   //__________________________________________________________________
   // Shotcounter mixinghead 08:
   //
         A     "DB619_State_MPart".Mixinghead[1].Shotcounter."08";
         =     "DB123_MH_IO_Signals".MH[8].OUT.MH.H_Shotcounter_MH;
         JCN   countMH8end;
   //
         A     "DB619_State_MPart".Mixinghead[1].ImpCounterOn;
         JCN   countMH8end;
   //-----
         L     "DB_Zaehler_Anzeige".MH_Counter_Reset[8];
         L     "DB619_State_MPart".Mixinghead[1].Countervalue;
         DTR;
         +R;
         T     "DB_Zaehler_Anzeige".MH_Counter_Reset[8];
   //-----
         L     "DB_Zaehler_Anzeige".MH_Counter_NonReset[8];
         L     "DB619_State_MPart".Mixinghead[1].Countervalue;
         DTR;
         +R;
         T     "DB_Zaehler_Anzeige".MH_Counter_NonReset[8];
   //-----
         L     "DB_Zaehler_Schicht_aktuell".MH_Counter[8];
         L     1.0;
         +R;
         T     "DB_Zaehler_Schicht_aktuell".MH_Counter[8];
   //-----
   countMH8end:NOP   0;
   //__________________________________________________________________
   // Shotcounter mixinghead 09:
   //
         A     "DB619_State_MPart".Mixinghead[1].Shotcounter."09";
         =     "DB123_MH_IO_Signals".MH[9].OUT.MH.H_Shotcounter_MH;
         JCN   countMH9end;
   //
         A     "DB619_State_MPart".Mixinghead[1].ImpCounterOn;
         JCN   countMH9end;
   //-----
         L     "DB_Zaehler_Anzeige".MH_Counter_Reset[9];
         L     "DB619_State_MPart".Mixinghead[1].Countervalue;
         DTR;
         +R;
         T     "DB_Zaehler_Anzeige".MH_Counter_Reset[9];
   //-----
         L     "DB_Zaehler_Anzeige".MH_Counter_NonReset[9];
         L     "DB619_State_MPart".Mixinghead[1].Countervalue;
         DTR;
         +R;
         T     "DB_Zaehler_Anzeige".MH_Counter_NonReset[9];
   //-----
         L     "DB_Zaehler_Schicht_aktuell".MH_Counter[9];
         L     1.0;
         +R;
         T     "DB_Zaehler_Schicht_aktuell".MH_Counter[9];
   //-----
   countMH9end:NOP   0;
   //__________________________________________________________________
   // Shotcounter mixinghead 10:
   //
         A     "DB619_State_MPart".Mixinghead[1].Shotcounter."10";
         =     "DB123_MH_IO_Signals".MH[10].OUT.MH.H_Shotcounter_MH;
         JCN   countMH10end;
   //
         A     "DB619_State_MPart".Mixinghead[1].ImpCounterOn;
         JCN   countMH10end;
   //-----
         L     "DB_Zaehler_Anzeige".MH_Counter_Reset[10];
         L     "DB619_State_MPart".Mixinghead[1].Countervalue;
         DTR;
         +R;
         T     "DB_Zaehler_Anzeige".MH_Counter_Reset[10];
   //-----
         L     "DB_Zaehler_Anzeige".MH_Counter_NonReset[10];
         L     "DB619_State_MPart".Mixinghead[1].Countervalue;
         DTR;
         +R;
         T     "DB_Zaehler_Anzeige".MH_Counter_NonReset[10];
   //-----
         L     "DB_Zaehler_Schicht_aktuell".MH_Counter[10];
         L     1.0;
         +R;
         T     "DB_Zaehler_Schicht_aktuell".MH_Counter[10];
   //-----
   countMH10end:NOP   0;
END_REGION

REGION Network 8: Bits for nozzle/bypass control on mixinghead
         BEU;
   //______________________________________________________________
   // send nozzles for shot from shot data
         L;
         LAR1;
         L     "DB619_State_MPart".ShotMa[1].ShotData.Comp_at_Shot;
         T     LB[AR1, P#0.0];

         L;
         LAR1;
         L     "DB704_MH_Value".Mixinghead[1].NozzelCirc;
         T     LB[AR1, P#0.0];

         A     #TempNozzleShotConnection[1];
         AN    "DB753_MeteringPump".Pump[1].PumpDeselected;
         AN    "DB753_MeteringPump".Pump[1].PumpDeselectedInterval;
         =     #TempNozzleShotMH[1];
         =     #TempNozzleCirc[1];
         A     #TempNozzleShotConnection[2];
         AN    "DB753_MeteringPump".Pump[2].PumpDeselected;
         AN    "DB753_MeteringPump".Pump[2].PumpDeselectedInterval;
         =     #TempNozzleShotMH[2];
         =     #TempNozzleCirc[2];
         A     #TempNozzleShotConnection[3];
         AN    "DB753_MeteringPump".Pump[3].PumpDeselected;
         AN    "DB753_MeteringPump".Pump[3].PumpDeselectedInterval;
         =     #TempNozzleShotMH[3];
         =     #TempNozzleCirc[3];
         A     #TempNozzleShotConnection[4];
         AN    "DB753_MeteringPump".Pump[4].PumpDeselected;
         AN    "DB753_MeteringPump".Pump[4].PumpDeselectedInterval;
         =     #TempNozzleShotMH[4];
         =     #TempNozzleCirc[4];

         CLR;
         =     #TempNozzleShotMH[5];
         =     #TempNozzleCirc[5];

         L;
         LAR1;
         L     LB[AR1, P#0.0];
         T     "DB704_MH_Value".Mixinghead[1].NozzelShot;

   //______________________________________________________________
   // Nozzles in recirculation are different between cycle and recirculation
         AN    "DB619_State_MPart".Cycle[1].running;
         JC    rec;
         A     "DB619_State_MPart".Cycle[1].StandByTimeRuns;
         A     "DB619_State_MPart".Cycle[1].LastShotinToolFinished;
         AN    "DB619_State_MPart".ToolMa[1].ShotFound;
         AN    "DB619_State_MPart".Cycle[1].PulsShotend;
         S     #TempNozzleCirc[1];
         S     #TempNozzleCirc[2];
         S     #TempNozzleCirc[3];
         S     #TempNozzleCirc[4];
         JU    orec;
   rec:  A     "DB619_State_MPart".Recirculation[1].Lowpressure;
         JC    lopr;
         A     "DB619_State_MPart".Recirculation[1].Reduced;
         JC    rdpr;
         A     "DB619_State_MPart".Recirculation[1].Highpressure;
         JC    hdpr;
         JU    orec;

   // nozzles for lo pressure recirculation
   lopr: NOP   0;
         A     "DB704_MH_Value".Mixinghead[1].MH_Connection[1].LP_CircOverNozzle;
         =     #TempNozzleCirc[1];
         A     "DB704_MH_Value".Mixinghead[1].MH_Connection[2].LP_CircOverNozzle;
         =     #TempNozzleCirc[2];
         A     "DB704_MH_Value".Mixinghead[1].MH_Connection[3].LP_CircOverNozzle;
         =     #TempNozzleCirc[3];
         A     "DB704_MH_Value".Mixinghead[1].MH_Connection[4].LP_CircOverNozzle;
         =     #TempNozzleCirc[4];
         JU    orec;
   // nozzles for reduced recirculation
   rdpr: A     "DB704_MH_Value".Mixinghead[1].MH_Connection[1].Red_CircOverNozzle;
         =     #TempNozzleCirc[1];
         A     "DB704_MH_Value".Mixinghead[1].MH_Connection[2].Red_CircOverNozzle;
         =     #TempNozzleCirc[2];
         A     "DB704_MH_Value".Mixinghead[1].MH_Connection[3].Red_CircOverNozzle;
         =     #TempNozzleCirc[3];
         A     "DB704_MH_Value".Mixinghead[1].MH_Connection[4].Red_CircOverNozzle;
         =     #TempNozzleCirc[4];
         JU    orec;
   // nozzles for high pressure recirculation
   hdpr: A     "DB704_MH_Value".Mixinghead[1].MH_Connection[1].HP_CircOverNozzle;
         =     #TempNozzleCirc[1];
         A     "DB704_MH_Value".Mixinghead[1].MH_Connection[2].HP_CircOverNozzle;
         =     #TempNozzleCirc[2];
         A     "DB704_MH_Value".Mixinghead[1].MH_Connection[3].HP_CircOverNozzle;
         =     #TempNozzleCirc[3];
         A     "DB704_MH_Value".Mixinghead[1].MH_Connection[4].HP_CircOverNozzle;
         =     #TempNozzleCirc[4];
         JU    orec;

   // switch deselected components to bypass before sending info to procan module
   orec: NOP   0;
         O     "DB753_MeteringPump".Pump[1].PumpDeselected;
         O     "DB613_Komponent_State".MeteringPump[1].IntervalPause;
         R     #TempNozzleCirc[1];
         O     "DB753_MeteringPump".Pump[2].PumpDeselected;
         O     "DB613_Komponent_State".MeteringPump[2].IntervalPause;
         R     #TempNozzleCirc[2];
         O     "DB753_MeteringPump".Pump[3].PumpDeselected;
         O     "DB613_Komponent_State".MeteringPump[3].IntervalPause;
         R     #TempNozzleCirc[3];
         O     "DB753_MeteringPump".Pump[4].PumpDeselected;
         O     "DB613_Komponent_State".MeteringPump[4].IntervalPause;
         R     #TempNozzleCirc[4];

         A     "TM_SwitchOnDelayFCPump";
         JCN   PUND;
         SET;
         R     #TempNozzleCirc[1];
         R     #TempNozzleCirc[2];
         R     #TempNozzleCirc[3];
         R     #TempNozzleCirc[4];
         JU    NozC;

   PUND: O     "DB619_State_MPart".Recirculation[1].Lowpressure;
         O     "DB619_State_MPart".Recirculation[1].Reduced;
         AN    "DB619_State_MPart".Recirculation[1].Pausetime;
         O     "DB619_State_MPart".Recirculation[1].Highpressure;
         O     "DB619_State_MPart".Cycle[1].running;
         JCN   mask;

   NozC: NOP   0;

         L;
         LAR1;
         L     LB[AR1, P#0.0];
         T     "DB704_MH_Value".Mixinghead[1].NozzelCirc;

   //______________________________________________________________
   // Mask with enable bits for the nozzle/bypass pairs
   mask: L;
         LAR1;
         L     0;
         T     LW[AR1, P#0.0];

   // Jump over enabling of nozzles when nozzle leakage test is active
         A     "DB704_MH_Value".Mixinghead[1].NozzleLeakageTest;
         A     "DB619_State_MPart".Operationmode[1].Manual;
         JC    test;

         A     "DB613_Komponent_State".MeteringPump[1].Main_Pumpselection;
         =     #TempMask.EnableNozzle_1;
         A     "DB613_Komponent_State".MeteringPump[2].Main_Pumpselection;
         =     #TempMask.EnableNozzle_2;
         A     "DB613_Komponent_State".MeteringPump[3].Main_Pumpselection;
         =     #TempMask.EnableNozzle_3;
         A     "DB613_Komponent_State".MeteringPump[4].Main_Pumpselection;
         =     #TempMask.EnableNozzle_4;

   test: L;
         LAR1;

         L     LW[AR1, P#0.0];  // target status
         L     "DB704_MH_Value".Mixinghead[1].NozzelForcen;  // old status
         XOW;  //  -> bits with differences
         AW;  // compare again with accu 2 -> bits to be switched on
         T     #SwitchOn;

         L     "DB704_MH_Value".Mixinghead[1].NozzelForcen;  // old status
         L     LW[AR1, P#0.0];  // target status
         XOW;  // -> bits with differences
         AW;  // compare again with accu 2 -> bits to be switched off
         T     #SwitchOff;

         A     <>0;
         L     "DB704_MH_Value".Mixinghead[1].DelayTimeNozzlesOff;
         SD    "TM_Nozzle_off_delay_MH01";
         A     "TM_Nozzle_off_delay_MH01";
         JCN   nzon;
         L     "DB704_MH_Value".Mixinghead[1].NozzelForcen;
         L     #SwitchOff;
         XOW;
         T     "DB704_MH_Value".Mixinghead[1].NozzelForcen;

   nzon: L     #SwitchOn;
         L     "DB704_MH_Value".Mixinghead[1].NozzelForcen;
         OW;
         T     "DB704_MH_Value".Mixinghead[1].NozzelForcen;

         A     "DB704_MH_Value".Mixinghead[1].NozzleLeakageTest;
         =     "DB824_Error_MH_CP".MH_Control[0].WRN_NozzleLeakageTest_active;
END_REGION
END_FUNCTION_BLOCK

FUNCTION_BLOCK "FB015_MeteringPump_M1"   // FB15, STL
TITLE = Meteringunit, edge filter, feed pump
{ S7_Optimized_Access := 'FALSE' }
AUTHOR : KT242
VERSION : 0.1
// Control of metering unit
   VAR_TEMP
      Dummy : Bool;
      Release_external : Bool;
      Release_FU : Bool;
      active : Bool;
      High_speed : Bool;
      V_2_Point_adjustment : Bool;
      Imp_WT_Ein : Bool;
      Imp_WT_Aus : Bool;
      HM_Intervall_Aus : Bool;
      Temp_F_FU_Poly : Bool;
      Temp_F_FU_Iso : Bool;
      Temp_enableCL_k1 : Bool;
      Temp_enableCL_k2 : Bool;
      Temp_Enable_C1 : Bool;
      Temp_Press_OK : Bool;
      CompUsedForShot : Array[1..16] of Bool;
      RetValSFC : Int;
   END_VAR
BEGIN

REGION Network 1: Min.- and Max.-value pump

         CALL  "FC217_Calc_flow_limits";
END_REGION

REGION Network 2

         CALL  "FC051_ComponentGeneral";
END_REGION

REGION Network 3: Temperautre control

         CALL  "FC057_HPHeatexchanger";
         CALL  "FC057_LPHeatexchanger";
END_REGION

REGION Network 4: Switch ON delay FU pump
   //-----
         O(;
         AN    "DB619_State_MPart".Machine[1].Metering."01";
         AN    "DB753_MeteringPump".Pump[1].PumpDeselected;
         A     "DB753_MeteringPump".Pump[1].WithFC;
         );
         O(;
         AN    "DB619_State_MPart".Machine[1].Metering."02";
         AN    "DB753_MeteringPump".Pump[2].PumpDeselected;
         A     "DB753_MeteringPump".Pump[2].WithFC;
         );
         O(;
         AN    "DB619_State_MPart".Machine[1].Metering."03";
         AN    "DB753_MeteringPump".Pump[3].PumpDeselected;
         A     "DB753_MeteringPump".Pump[3].WithFC;
         );
         O(;
         AN    "DB619_State_MPart".Machine[1].Metering."04";
         AN    "DB753_MeteringPump".Pump[4].PumpDeselected;
         A     "DB753_MeteringPump".Pump[4].WithFC;
         );
         O(;
         AN    "DB619_State_MPart".Machine[1].Metering."05";
         AN    "DB753_MeteringPump".Pump[5].PumpDeselected;
         A     "DB753_MeteringPump".Pump[5].WithFC;
         );
         O(;
         AN    "DB619_State_MPart".Machine[1].Metering."06";
         AN    "DB753_MeteringPump".Pump[6].PumpDeselected;
         A     "DB753_MeteringPump".Pump[6].WithFC;
         );
         FP    "HF_FP_SwitchOffPump";
         =     "PulsePumpSwitchedOff";
         L     S5T#5S;
         SE    "TM_SwitchOnDelayFCPump";
   //-----
END_REGION

REGION Network 5: Release of pumps
   // Copy Control bits for module to local area
         L;
         LAR1;
         L     "DB619_State_MPart".ShotMa[1].ShotData.Comp_at_Shot;
         CAW;
         T     LW[AR1, P#0.0];
   //-----
         A(;
         O     "DB619_State_MPart".CylinderManager[1].Selection_Metering;
         ON    "DB619_State_MPart".CylinderManager[1].Block_is_active;
         );
   //-----
         A(;
         O     "DB613_Komponent_State".MeteringPump[1].Main_Pumpselection;
         O     "DB753_MeteringPump".Pump[1].PumpDeselected;
         O     "DB613_Komponent_State".MeteringPump[1].IntervalPause;
         ON    "DB613_Komponent_State".MeteringPump[1].Block_is_active;
         );
         A(;
         O     "DB613_Komponent_State".MeteringPump[2].Main_Pumpselection;
         O     "DB753_MeteringPump".Pump[2].PumpDeselected;
         O     "DB613_Komponent_State".MeteringPump[2].IntervalPause;
         ON    "DB613_Komponent_State".MeteringPump[2].Block_is_active;
         );
         A(;
         O     "DB613_Komponent_State".MeteringPump[3].Main_Pumpselection;
         O     "DB753_MeteringPump".Pump[3].PumpDeselected;
         O     "DB613_Komponent_State".MeteringPump[3].IntervalPause;
         ON    "DB613_Komponent_State".MeteringPump[3].Block_is_active;
         );
         A(;
         O     "DB613_Komponent_State".MeteringPump[4].Main_Pumpselection;
         O     "DB753_MeteringPump".Pump[4].PumpDeselected;
         O     "DB613_Komponent_State".MeteringPump[4].IntervalPause;
         ON    "DB613_Komponent_State".MeteringPump[4].Block_is_active;
         );
         A(;
         O     "DB613_Komponent_State".MeteringPump[5].Main_Pumpselection;
         O     "DB753_MeteringPump".Pump[5].PumpDeselected;
         O     "DB613_Komponent_State".MeteringPump[5].IntervalPause;
         ON    "DB613_Komponent_State".MeteringPump[5].Block_is_active;
         );
         A(;
         O     "DB613_Komponent_State".MeteringPump[6].Main_Pumpselection;
         O     "DB753_MeteringPump".Pump[6].PumpDeselected;
         O     "DB613_Komponent_State".MeteringPump[6].IntervalPause;
         ON    "DB613_Komponent_State".MeteringPump[6].Block_is_active;
         );
         AN    "TM_SwitchOnDelayFCPump";
         AN    "TM_Interrupt2PointAdjustment";
         =     #Release_external;
   //-----
END_REGION

REGION Network 6: Preparation for 2 Point- Adjustment
         CALL  "FC216_2-point_adjust";
END_REGION

REGION Network 7: Component 1
   //___________________________________________________________________________
   // Feedpump component 1
   //___________________________________________________________________________
   //
         CALL  "FC123_FeedingPump"
         ( IN_Release               := "DB619_State_MPart".Operationmode[1].valid,
           IN_ControlVoltage        := "DB619_State_MPart".Operationmode[1].Controllvoltage,
           IN_Reset_fault           := "DB009_Faults".Faults_Reset_FKT_M1,
           IN_ComponentDeselected   := "DB613_Komponent_State".MeteringPump[1].Mes_PumpDeselected,
           IN_Request_Feed          := "DB613_Komponent_State".MeteringPump[1].Selection_Feedingpump,
           IN_Request_Filling       := "DB612_Tank_State".Tank[1].Filling_Start,
           IN_Request_Bypass        := 1,
           IN_Fault_Motorprotection := "F_FeedingP_C1",
           IN_FaultFreqConverter    := "F_FCFeedingP_C1",
           IN_DryRun                := "DB612_Tank_State".Tank[1].Min_Level,
           IN_MaxLevelTray          := "DB612_Tank_State".Tank[1].LevelTriptray,
           IN_MaxPressure           := 1,
           IN_TempRelease           := 1,
           IN_TimerDrive            := "TM1_FeedPump01",
           IN_TimerStartUpFConv     := "TM2_FeedPump01",
           Values                   := "DB751_auxiliaryDriveMetering".FeedingPump[1],
           OUT_MainsContactor       := "M_FeedingP_C1",
           OUT_Release_FConverter   := "M_FeedingP_Start_C1",
           IO_Status                := "DB613_Komponent_State".FeedPump[1],
           IO_NewFault              := "DB009_Faults".Faultschanging_M1,
           IO_FaultLevel_1          := "DB009_Faults".Faults_FKT_Grp_1_M1,
           IO_FaultLevel_3          := "DB009_Faults".Faults_FKT_Grp_3_M1,
           IO_Faults                := "DB823_Error_Metering".FeedPump[1]
         );
   //___________________________________________________________________________
   // Edgefilter component 1
   //___________________________________________________________________________
   //
         CALL  "FC122_EdgeFilter"
         ( IN_Release               := "DB619_State_MPart".Operationmode[1].valid,
           IN_Reset_fault           := "DB009_Faults".Faults_Reset_FKT_M1,
           IN_Fault_Motorprotection := "F_Platefilter_C1",
           IN_DifPressure           := FALSE,
           IN_TimerDrive            := "TM_EdgeFilter01",
           Values                   := "DB751_auxiliaryDriveMetering".EdgeFilter[1],
           OUT_MainsContactor       := "M_Platefilter_C1",
           IO_Status                := "DB613_Komponent_State".EdgeFilter[1],
           IO_NewFault              := "DB009_Faults".Faultschanging_M1,
           IO_FaultLevel_3          := "DB009_Faults".Faults_FKT_Grp_3_M1,
           IO_Faults                := "DB823_Error_Metering".EdgeFilter[1]
         );
   //___________________________________________________________________________
   // Metering pump component 1
   //___________________________________________________________________________
   //
         A     "P_Min_C1";
         O;
         A     "DB619_State_MPart".Operationmode[1].Test;
         A     "V_Bypass_C1";
         =     #Temp_Press_OK;

         O     "DB612_Tank_State".Pentan[1].EnableComponentPump;
         ON    "DB702_Tank_Value".Tank[1].With_Filling_Pentane;
         A     #Release_external;
         =     #Temp_Enable_C1;
   //-----
         CALL  "FC053_MeteringPump"
         ( IN_ControlVoltage        := "DB619_State_MPart".Operationmode[1].Controllvoltage,
           IN_OperationMode_Valid   := #Release_external,
           IN_OPerationMode_Active  := "DB619_State_MPart".Operationmode[1].Active,
           IN_Min_PrePressure       := "P_Prepressure_Pump_C1",
           IN_Max_PressureComponent := "P_Max_C1",
           IN_MotorprotectionPump   := "F_Pump_C1",
           IN_With_FU_Pump          := "DB753_MeteringPump".Pump[1].WithFC,
           IN_FLT_FU_Pump           := "F_FC_Pump_C1",
           IN_MaxLevelTray          := "L_DripTray_C1",
           IN_Shot_Start            := "DB619_State_MPart".Cycle[1].Shotrelease,
           IN_MinPressure           := #Temp_Press_OK,  //"P_Min_C1"
           IN_PreAlarmBearing       := FALSE,  // "F_PreAlarmBearing_K2"
           IN_AlarmBearing          := FALSE,  // "F_AlarmBearing_K2"
           IN_Reset_fault_Fkt       := "DB009_Faults".Faults_Reset_FKT_M1,
           IN_ReleaseExternal       := #Temp_Enable_C1,  // #Release_external
           IN_FaultGroup_1          := "DB009_Faults".Fault_State_Grp_1_M1,
           IN_SOverSOffSWU_running  := "DB619_State_MPart".SWU[1].Switchingtime_runs,
           IN_High_speed            := 0,
           IN_2point_Adjustment     := "DB613_Komponent_State".MeteringPump[1]."2PointAdjustmentSelected",
           IN_Cycle_running         := "DB619_State_MPart".Cycle[1].running,
           IN_Recirc_reduced        := "DB619_State_MPart".Recirculation[1].Reduced,
           IN_Recirc_lowpressure    := "DB619_State_MPart".Recirculation[1].Lowpressure,
           IN_Recirc_highpressure   := "DB619_State_MPart".Recirculation[1].Highpressure,
           IN_Recirc_pausetime      := "DB619_State_MPart".Recirculation[1].Pausetime,
           IN_UsedForShot           := #CompUsedForShot[1],
           IN_Delay_Restart         := S5T#2S,
           IN_Timer_Restart         := "TM_RestartC01",
           IN_RunDownTime_FeedPump  := S5T#3S,
           IN_Timer_ControlFeedPump := "TM_CtrlFeedPumpC01",
           IN_TimerOffFeedPump      := "TM_CommonC01",
           IN_Timer_Delay_EnClosedL := "TM_DelayClosedLoopC01",
           IN_TimerInterval         := "TM_IntervalC01",
           OUT_2_Point_Adjust       := #V_2_Point_adjustment,
           OUT_Dosing_active        := #Dummy,
           OUT_Enableclosedloop     := "DB122_FlowIndexState".MeteringUnit[1].OUT_PROCAN.FlowIndex.Enableclosedloop,
           OUT_Pump_MainsContactor  := "M_Pump_Net_C1",
           OUT_Release_FU           := "M_Pump_Start_C1",
           IO_QPB_Pumpe             := "DB122_FlowIndexState".MeteringUnit[1].OUT_PROCAN.FlowIndex.StartQPB,
           IO_Status                := "DB613_Komponent_State".MeteringPump[1],
           IO_Fault                 := "DB823_Error_Metering".MeteringPump[1],
           IO_Config                := "DB753_MeteringPump".Pump[1],
           IO_NewFault              := "DB009_Faults".Faultschanging_M1,
           IO_FaultLevel_1          := "DB009_Faults".Faults_FKT_Grp_1_M1,
           IO_FaultLevel_2          := "DB009_Faults".Faults_FKT_Grp_2_M1,
           IO_FaultLevel_3          := "DB009_Faults".Faults_FKT_Grp_3_M1
         );
   //-----
   //-----
   // 2 Point adjustment
         A     #V_2_Point_adjustment;
         L     s5t#800ms;
         SE    "TM_pulse_2PointAdjust_C1";

         A     #V_2_Point_adjustment;
         L     s5t#500ms;
         SD    "TM_delay_2PointAdjust_C1";
         A     "TM_delay_2PointAdjust_C1";
         =     "V_Pump_2Point_C1";
   //-----
   //
         A     "DB613_Komponent_State".MeteringPump[1].Metering_to_PUC;
         =     "DB619_State_MPart".Machine[1].Metering."01";
   //
         A     "DB613_Komponent_State".MeteringPump[1].Metering_to_PUC;
         =     "M1C01active";
   //___________________________________________________________________________
   // Ventilation metering pump component 1
   //___________________________________________________________________________
   //
         CALL  "FC055_PumpVentilation"
         ( IN_Reset_fault_Fkt     := "DB009_Faults".Faults_Reset_FKT_M1,
           IN_Motorprotection     := "F_Fan_Pump_C1",
           IN_ComponentDeselected := "DB613_Komponent_State".MeteringPump[1].Mes_PumpDeselected,
           In_Start               := "DB613_Komponent_State".MeteringPump[1].Metering_to_PUC,
           IN_Time                := S5T#1M,
           IN_Timer               := "TM_FanPumpC01",
           OUT_MainContactor      := "M_Fan_Pump_Net_C1",
           IO_FLT_MotorFan        := "DB823_Error_Metering".MeteringPump[1].FLT_MotorFan,
           IO_NewFault            := "DB009_Faults".Faultschanging_M1,
           IO_FaultLevel_2        := "DB009_Faults".Faults_FKT_Grp_2_M1,
           IO_FaultLevel_3        := "DB009_Faults".Faults_FKT_Grp_3_M1
         );
   //
END_REGION

REGION Network 8: Component 2
   //___________________________________________________________________________
   // Feedpump component 2
   //___________________________________________________________________________
   //
         CALL  "FC123_FeedingPump"
         ( IN_Release               := "DB619_State_MPart".Operationmode[1].valid,
           IN_ControlVoltage        := "DB619_State_MPart".Operationmode[1].Controllvoltage,
           IN_Reset_fault           := "DB009_Faults".Faults_Reset_FKT_M1,
           IN_ComponentDeselected   := "DB613_Komponent_State".MeteringPump[2].Mes_PumpDeselected,
           IN_Request_Feed          := "DB613_Komponent_State".MeteringPump[2].Selection_Feedingpump,
           IN_Request_Filling       := 0,
           IN_Request_Bypass        := 0,
           IN_Fault_Motorprotection := "F_FeedingP_C2",
           IN_FaultFreqConverter    := "F_FCFeedingP_C2",
           IN_DryRun                := "DB612_Tank_State".Tank[2].Min_Level,
           IN_MaxLevelTray          := "DB612_Tank_State".Tank[2].LevelTriptray,
           IN_MaxPressure           := 1,
           IN_TempRelease           := 1,
           IN_TimerDrive            := "TM1_FeedPump02",
           IN_TimerStartUpFConv     := "TM2_FeedPump02",
           Values                   := "DB751_auxiliaryDriveMetering".FeedingPump[2],
           OUT_MainsContactor       := "M_FeedingP_C2",
           OUT_Release_FConverter   := "M_FeedingP_Start_C2",
           IO_Status                := "DB613_Komponent_State".FeedPump[2],
           IO_NewFault              := "DB009_Faults".Faultschanging_M1,
           IO_FaultLevel_1          := "DB009_Faults".Faults_FKT_Grp_1_M1,
           IO_FaultLevel_3          := "DB009_Faults".Faults_FKT_Grp_3_M1,
           IO_Faults                := "DB823_Error_Metering".FeedPump[2]
         );
   //___________________________________________________________________________
   // Edgefilter component 2
   //___________________________________________________________________________
   //
         CALL  "FC122_EdgeFilter"
         ( IN_Release               := "DB619_State_MPart".Operationmode[1].valid,
           IN_Reset_fault           := "DB009_Faults".Faults_Reset_FKT_M1,
           IN_Fault_Motorprotection := "F_Platefilter_C2",
           IN_DifPressure           := FALSE,
           IN_TimerDrive            := "TM_EdgeFilter02",
           Values                   := "DB751_auxiliaryDriveMetering".EdgeFilter[2],
           OUT_MainsContactor       := "M_Platefilter_C2",
           IO_Status                := "DB613_Komponent_State".EdgeFilter[2],
           IO_NewFault              := "DB009_Faults".Faultschanging_M1,
           IO_FaultLevel_3          := "DB009_Faults".Faults_FKT_Grp_3_M1,
           IO_Faults                := "DB823_Error_Metering".EdgeFilter[2]
         );
   //___________________________________________________________________________
   // Metering pump component 2
   //___________________________________________________________________________
   //
         A     "P_Min_C2";
         O;
         A     "DB619_State_MPart".Operationmode[1].Test;
         A     "V_Bypass_C2";
         =     #Temp_Press_OK;

         CALL  "FC053_MeteringPump"
         ( IN_ControlVoltage        := "DB619_State_MPart".Operationmode[1].Controllvoltage,
           IN_OperationMode_Valid   := #Release_external,  // not used at FC
           IN_OPerationMode_Active  := "DB619_State_MPart".Operationmode[1].Active,
           IN_Min_PrePressure       := "P_Prepressure_Pump_C2",
           IN_Max_PressureComponent := "P_Max_C2",
           IN_MotorprotectionPump   := "F_Pump_C2",
           IN_With_FU_Pump          := "DB753_MeteringPump".Pump[2].WithFC,
           IN_FLT_FU_Pump           := "F_FC_Pump_C2",
           IN_MaxLevelTray          := "L_DripTray_C2",
           IN_Shot_Start            := "DB619_State_MPart".Cycle[1].Shotrelease,
           IN_MinPressure           := #Temp_Press_OK,  //"P_Min_C2"
           IN_PreAlarmBearing       := FALSE,  // "F_PreAlarmBearing_K2"
           IN_AlarmBearing          := FALSE,  // "F_AlarmBearing_K2"
           IN_Reset_fault_Fkt       := "DB009_Faults".Faults_Reset_FKT_M1,
           IN_ReleaseExternal       := #Release_external,
           IN_FaultGroup_1          := "DB009_Faults".Fault_State_Grp_1_M1,
           IN_SOverSOffSWU_running  := "DB619_State_MPart".SWU[1].Switchingtime_runs,
           IN_High_speed            := 0,
           IN_2point_Adjustment     := "DB613_Komponent_State".MeteringPump[2]."2PointAdjustmentSelected",
           IN_Cycle_running         := "DB619_State_MPart".Cycle[1].running,
           IN_Recirc_reduced        := "DB619_State_MPart".Recirculation[1].Reduced,
           IN_Recirc_lowpressure    := "DB619_State_MPart".Recirculation[1].Lowpressure,
           IN_Recirc_highpressure   := "DB619_State_MPart".Recirculation[1].Highpressure,
           IN_Recirc_pausetime      := "DB619_State_MPart".Recirculation[1].Pausetime,
           IN_UsedForShot           := #CompUsedForShot[2],
           IN_Delay_Restart         := S5T#2S,
           IN_Timer_Restart         := "TM_RestartC02",
           IN_RunDownTime_FeedPump  := S5T#3S,
           IN_Timer_ControlFeedPump := "TM_CtrlFeedPumpC02",
           IN_TimerOffFeedPump      := "TM_CommonC02",
           IN_Timer_Delay_EnClosedL := "TM_DelayClosedLoopC02",
           IN_TimerInterval         := "TM_IntervalC02",
           OUT_2_Point_Adjust       := #V_2_Point_adjustment,
           OUT_Dosing_active        := #Dummy,
           OUT_Enableclosedloop     := "DB122_FlowIndexState".MeteringUnit[2].OUT_PROCAN.FlowIndex.Enableclosedloop,
           OUT_Pump_MainsContactor  := "M_Pump_Net_C2",
           OUT_Release_FU           := "M_Pump_Start_C2",
           IO_QPB_Pumpe             := "DB122_FlowIndexState".MeteringUnit[2].OUT_PROCAN.FlowIndex.StartQPB,
           IO_Status                := "DB613_Komponent_State".MeteringPump[2],
           IO_Fault                 := "DB823_Error_Metering".MeteringPump[2],
           IO_Config                := "DB753_MeteringPump".Pump[2],
           IO_NewFault              := "DB009_Faults".Faultschanging_M1,
           IO_FaultLevel_1          := "DB009_Faults".Faults_FKT_Grp_1_M1,
           IO_FaultLevel_2          := "DB009_Faults".Faults_FKT_Grp_2_M1,
           IO_FaultLevel_3          := "DB009_Faults".Faults_FKT_Grp_3_M1
         );
   //-----
   // 2 Point adjustment
         A     #V_2_Point_adjustment;
         L     s5t#800ms;
         SE    "TM_pulse_2PointAdjust_C2";

         A     #V_2_Point_adjustment;
         L     s5t#500ms;
         SD    "TM_delay_2PointAdjust_C2";
         A     "TM_delay_2PointAdjust_C2";
         =     "V_Pump_2Point_C2";
   //-----
   //
         A     "DB613_Komponent_State".MeteringPump[2].Metering_to_PUC;
         =     "DB619_State_MPart".Machine[1].Metering."02";
   //
         A     "DB613_Komponent_State".MeteringPump[2].Metering_to_PUC;
         =     "M1C02active";
   //___________________________________________________________________________
   // Ventilation metering pump component 2
   //___________________________________________________________________________
   //
         CALL  "FC055_PumpVentilation"
         ( IN_Reset_fault_Fkt     := "DB009_Faults".Faults_Reset_FKT_M1,
           IN_Motorprotection     := "F_Fan_Pump_C2",
           IN_ComponentDeselected := "DB613_Komponent_State".MeteringPump[2].Mes_PumpDeselected,
           In_Start               := "DB613_Komponent_State".MeteringPump[2].Metering_to_PUC,
           IN_Time                := S5T#1M,
           IN_Timer               := "TM_FanPumpC02",
           OUT_MainContactor      := "M_Fan_Pump_Net_C2",
           IO_FLT_MotorFan        := "DB823_Error_Metering".MeteringPump[2].FLT_MotorFan,
           IO_NewFault            := "DB009_Faults".Faultschanging_M1,
           IO_FaultLevel_2        := "DB009_Faults".Faults_FKT_Grp_2_M1,
           IO_FaultLevel_3        := "DB009_Faults".Faults_FKT_Grp_3_M1
         );
   //-----
END_REGION
END_FUNCTION_BLOCK

FUNCTION_BLOCK "FB017_CPiston_M1"   // FB17, STL
TITLE = cleaning pistons of mixingheads
{ S7_Optimized_Access := 'FALSE' }
AUTHOR : KT242
VERSION : 0.1
// Activation of cleaning piston mixinghead
   VAR_TEMP
      RetValSFC : Int;
      AnaCp_Stat : Word;
      AnaCp_StatB : Byte;
      Temp_AnaCP : Bool;
      Temp_CP_forward_external : Bool;
      Temp_Shotend : Bool;
   END_VAR
BEGIN

REGION Network 1: Activate cleaning piston mixinghead by external signal
         A     "DB005_RS<->Extern".MC_Interface[1].Data_from_MC.CP_forward;
         O     "DB1900_IF_Robots".State_Robots[1].CleaningMHOn;
         O(;
         A     "DB2000_FRA<->KM".Input.comandstatus.CPFORWARD;
         A     "S_Automatic_MH01";
         );
         =     #Temp_CP_forward_external;
END_REGION

REGION Network 2: Cleaning piston mixinghead 01
         CALL  BLKMOV
         ( SRCBLK  := "DB123_MH_IO_Signals".MH[1].IN.CleaningPistonState,
           RET_VAL := #RetValSFC,
           DSTBLK  := #AnaCp_Stat
         );

         L     #AnaCp_Stat;
         SRW   8;
         T     #AnaCp_StatB;

         A     "DB619_State_MPart".Cycle[1].PulsShotend;
         O;
         A(;
         A     "DB123_MH_IO_Signals".MH[1].IN.MH_Aps_Mixinghead;
         A     "DB619_State_MPart".Operationmode[1].Test;
         FN    "HM_Shotend";
         );
         =     #Temp_Shotend;

         CALL  "FC071_CleaningPiston"
         ( IN_WithCP                := "DB704_MH_Value".Mixinghead[1].WithCleaningPiston,
           IN_Ana_CP_State          := #AnaCp_StatB,
           IN_SWUEnabled            := "DB619_State_MPart".SWU[1].SWU_released."01",
           IN_ButtonCPForward       := "DB123_MH_IO_Signals".MH[1].IN.MH_CP_forward,
           IN_ButtonCPback          := "DB123_MH_IO_Signals".MH[1].IN.MH_CP_backward,
           IN_CPForwardFromExternal := #Temp_CP_forward_external,
           IN_CPAfterShot           := "DB619_State_MPart".ShotMa[1].ShotData.CP_AfterShot,
           IN_PartshotDisabled      := "DB619_State_MPart".ShotMa[1].ShotData.ShotDisabled,
           IN_Blowing_OUT           := "DB614_MH_State".InertingMH[1].Start_Prepare_Purge_after_Shot,
           IN_CPProxSwitch          := "DB123_MH_IO_Signals".MH[1].IN.MH_APS_CleaningPiston,
           IN_SWUActive             := "DB619_State_MPart".SWU[1].Open_SWU_allone."01",
           IN_HydraulicOk           := "DB619_State_MPart".Machine[1].HydStartUp_finished,
           IN_ResetFaults           := "DB009_Faults".Faults_Reset_FKT_M1,
           IN_ControlVoltage        := "DB619_State_MPart".Operationmode[1].Controllvoltage,
           IN_OperatingModeValid    := "DB619_State_MPart".Operationmode[1].valid,
           IN_OperatingModeWithFoam := "DB619_State_MPart".Operationmode[1].Operation,
           IN_OperatingModeTestValv := FALSE,  //"DB619_State_MPart".Operationmode[1].Test
           IN_Lamptest              := "DB619_State_MPart".Operationmode[1].Lamptest,
           IN_ShotEnd               := #Temp_Shotend,
           IN_FaultLevel_1          := "DB009_Faults".Fault_State_Grp_1_M1,
           IN_PressurizeTimeRunning := "DB619_State_MPart".Cycle[1].PressurizeTimeRuns,
           IN_ShotActive            := "DB619_State_MPart".Cycle[1].ShotRuns,
           IN_CycleRunning          := "DB619_State_MPart".Cycle[1].running,
           IN_RmpCtrlChangeTimeEnd  := "DB619_State_MPart".Cycle[1].RmpCtrlChangeTimeEnd,
           IN_StandbyTimeRunning    := "DB619_State_MPart".Cycle[1].StandByTimeRuns,
           IN_RmpCycleEnd           := "DB619_State_MPart".Cycle[1].PulseCycleEnd,
           IN_CPTimer               := "TM_RunTime_CP01",
           IN_TMCheckHomePos        := "TM_FltCPHomePos_CP01",
           Values                   := "DB704_MH_Value".Mixinghead[1].Cleaning_Piston,
           OUT_ValveCPForward       := "DB123_MH_IO_Signals".MH[1].OUT.MH.V_CP_Forward_MH,
           OUT_LampCPBack           := "DB123_MH_IO_Signals".MH[1].OUT.MH.H_CP_Back_MH,
           IO_CPIsOk                := "DB619_State_MPart".Mixinghead[1].Cleaningpiston_OK,
           IO_ReqHydrForCleaning    := "DB611_Hydraulic_State".MH_Hydraulic[1].Request_from_CP,
           IO_Status                := "DB614_MH_State".MH_CleaningPiston[1],
           IO_Fault                 := "DB824_Error_MH_CP".CPiston[1],
           IO_NewFault              := "DB009_Faults".Faultschanging_M1,
           IO_FaultLevel_1          := "DB009_Faults".Faults_FKT_Grp_1_M1,
           IO_FaultLevel_2          := "DB009_Faults".Faults_FKT_Grp_2_M1,
           IO_FaultLevel_3          := "DB009_Faults".Faults_FKT_Grp_3_M1
         );
END_REGION

REGION Network 3: Activate cleaning piston mixinghead by external signal
         A     "DB005_RS<->Extern".MC_Interface[2].Data_from_MC.CP_forward;
         =     #Temp_CP_forward_external;
END_REGION

REGION Network 4: Cleaning piston mixinghead 02
         CALL  BLKMOV
         ( SRCBLK  := "DB123_MH_IO_Signals".MH[2].IN.CleaningPistonState,
           RET_VAL := #RetValSFC,
           DSTBLK  := #AnaCp_Stat
         );

         L     #AnaCp_Stat;
         SRW   8;
         T     #AnaCp_StatB;

         CALL  "FC071_CleaningPiston"
         ( IN_WithCP                := "DB704_MH_Value".Mixinghead[2].WithCleaningPiston,
           IN_Ana_CP_State          := #AnaCp_StatB,
           IN_SWUEnabled            := "DB619_State_MPart".SWU[1].SWU_released."02",
           IN_ButtonCPForward       := "DB123_MH_IO_Signals".MH[2].IN.MH_CP_forward,
           IN_ButtonCPback          := "DB123_MH_IO_Signals".MH[2].IN.MH_CP_backward,
           IN_CPForwardFromExternal := #Temp_CP_forward_external,
           IN_CPAfterShot           := "DB619_State_MPart".ShotMa[1].ShotData.CP_AfterShot,
           IN_PartshotDisabled      := "DB619_State_MPart".ShotMa[1].ShotData.ShotDisabled,
           IN_Blowing_OUT           := "DB614_MH_State".InertingMH[2].Start_Prepare_Purge_after_Shot,
           IN_CPProxSwitch          := "DB123_MH_IO_Signals".MH[2].IN.MH_APS_CleaningPiston,
           IN_SWUActive             := "DB619_State_MPart".SWU[1].Open_SWU_allone."02",
           IN_HydraulicOk           := "DB619_State_MPart".Machine[1].HydStartUp_finished,
           IN_ResetFaults           := "DB009_Faults".Faults_Reset_FKT_M1,
           IN_ControlVoltage        := "DB619_State_MPart".Operationmode[1].Controllvoltage,
           IN_OperatingModeValid    := "DB619_State_MPart".Operationmode[1].valid,
           IN_OperatingModeWithFoam := "DB619_State_MPart".Operationmode[1].Operation,
           IN_OperatingModeTestValv := "DB619_State_MPart".Operationmode[1].Test,
           IN_Lamptest              := "DB619_State_MPart".Operationmode[1].Lamptest,
           IN_ShotEnd               := "DB619_State_MPart".Cycle[1].PulsShotend,
           IN_FaultLevel_1          := "DB009_Faults".Fault_State_Grp_1_M1,
           IN_PressurizeTimeRunning := "DB619_State_MPart".Cycle[1].PressurizeTimeRuns,
           IN_ShotActive            := "DB619_State_MPart".Cycle[1].ShotRuns,
           IN_CycleRunning          := "DB619_State_MPart".Cycle[1].running,
           IN_RmpCtrlChangeTimeEnd  := "DB619_State_MPart".Cycle[1].RmpCtrlChangeTimeEnd,
           IN_StandbyTimeRunning    := "DB619_State_MPart".Cycle[1].StandByTimeRuns,
           IN_RmpCycleEnd           := "DB619_State_MPart".Cycle[1].PulseCycleEnd,
           IN_CPTimer               := "TM_RunTime_CP02",
           IN_TMCheckHomePos        := "TM_FltCPHomePos_CP02",
           Values                   := "DB704_MH_Value".Mixinghead[2].Cleaning_Piston,
           OUT_ValveCPForward       := "DB123_MH_IO_Signals".MH[2].OUT.MH.V_CP_Forward_MH,
           OUT_LampCPBack           := "DB123_MH_IO_Signals".MH[2].OUT.MH.H_CP_Back_MH,
           IO_CPIsOk                := "DB619_State_MPart".Mixinghead[1].Cleaningpiston_OK,
           IO_ReqHydrForCleaning    := "DB611_Hydraulic_State".MH_Hydraulic[1].Request_from_CP,
           IO_Status                := "DB614_MH_State".MH_CleaningPiston[2],
           IO_Fault                 := "DB824_Error_MH_CP".CPiston[2],
           IO_NewFault              := "DB009_Faults".Faultschanging_M1,
           IO_FaultLevel_1          := "DB009_Faults".Faults_FKT_Grp_1_M1,
           IO_FaultLevel_2          := "DB009_Faults".Faults_FKT_Grp_2_M1,
           IO_FaultLevel_3          := "DB009_Faults".Faults_FKT_Grp_3_M1
         );
END_REGION

REGION Network 5: Activate cleaning piston mixinghead by external signal
         A     "DB005_RS<->Extern".MC_Interface[3].Data_from_MC.CP_forward;
         =     #Temp_CP_forward_external;
END_REGION

REGION Network 6: Cleaning piston mixinghead 03
         CALL  BLKMOV
         ( SRCBLK  := "DB123_MH_IO_Signals".MH[3].IN.CleaningPistonState,
           RET_VAL := #RetValSFC,
           DSTBLK  := #AnaCp_Stat
         );

         L     #AnaCp_Stat;
         SRW   8;
         T     #AnaCp_StatB;

         CALL  "FC071_CleaningPiston"
         ( IN_WithCP                := "DB704_MH_Value".Mixinghead[3].WithCleaningPiston,
           IN_Ana_CP_State          := #AnaCp_StatB,
           IN_SWUEnabled            := "DB619_State_MPart".SWU[1].SWU_released."03",
           IN_ButtonCPForward       := "DB123_MH_IO_Signals".MH[3].IN.MH_CP_forward,
           IN_ButtonCPback          := "DB123_MH_IO_Signals".MH[3].IN.MH_CP_backward,
           IN_CPForwardFromExternal := #Temp_CP_forward_external,
           IN_CPAfterShot           := "DB619_State_MPart".ShotMa[1].ShotData.CP_AfterShot,
           IN_PartshotDisabled      := "DB619_State_MPart".ShotMa[1].ShotData.ShotDisabled,
           IN_Blowing_OUT           := "DB614_MH_State".InertingMH[3].Start_Prepare_Purge_after_Shot,
           IN_CPProxSwitch          := "DB123_MH_IO_Signals".MH[3].IN.MH_APS_CleaningPiston,
           IN_SWUActive             := "DB619_State_MPart".SWU[1].Open_SWU_allone."03",
           IN_HydraulicOk           := "DB619_State_MPart".Machine[1].HydStartUp_finished,
           IN_ResetFaults           := "DB009_Faults".Faults_Reset_FKT_M1,
           IN_ControlVoltage        := "DB619_State_MPart".Operationmode[1].Controllvoltage,
           IN_OperatingModeValid    := "DB619_State_MPart".Operationmode[1].valid,
           IN_OperatingModeWithFoam := "DB619_State_MPart".Operationmode[1].Operation,
           IN_OperatingModeTestValv := "DB619_State_MPart".Operationmode[1].Test,
           IN_Lamptest              := "DB619_State_MPart".Operationmode[1].Lamptest,
           IN_ShotEnd               := "DB619_State_MPart".Cycle[1].PulsShotend,
           IN_FaultLevel_1          := "DB009_Faults".Fault_State_Grp_1_M1,
           IN_PressurizeTimeRunning := "DB619_State_MPart".Cycle[1].PressurizeTimeRuns,
           IN_ShotActive            := "DB619_State_MPart".Cycle[1].ShotRuns,
           IN_CycleRunning          := "DB619_State_MPart".Cycle[1].running,
           IN_RmpCtrlChangeTimeEnd  := "DB619_State_MPart".Cycle[1].RmpCtrlChangeTimeEnd,
           IN_StandbyTimeRunning    := "DB619_State_MPart".Cycle[1].StandByTimeRuns,
           IN_RmpCycleEnd           := "DB619_State_MPart".Cycle[1].PulseCycleEnd,
           IN_CPTimer               := "TM_RunTime_CP03",
           IN_TMCheckHomePos        := "TM_FltCPHomePos_CP03",
           Values                   := "DB704_MH_Value".Mixinghead[3].Cleaning_Piston,
           OUT_ValveCPForward       := "DB123_MH_IO_Signals".MH[3].OUT.MH.V_CP_Forward_MH,
           OUT_LampCPBack           := "DB123_MH_IO_Signals".MH[3].OUT.MH.H_CP_Back_MH,
           IO_CPIsOk                := "DB619_State_MPart".Mixinghead[1].Cleaningpiston_OK,
           IO_ReqHydrForCleaning    := "DB611_Hydraulic_State".MH_Hydraulic[1].Request_from_CP,
           IO_Status                := "DB614_MH_State".MH_CleaningPiston[3],
           IO_Fault                 := "DB824_Error_MH_CP".CPiston[3],
           IO_NewFault              := "DB009_Faults".Faultschanging_M1,
           IO_FaultLevel_1          := "DB009_Faults".Faults_FKT_Grp_1_M1,
           IO_FaultLevel_2          := "DB009_Faults".Faults_FKT_Grp_2_M1,
           IO_FaultLevel_3          := "DB009_Faults".Faults_FKT_Grp_3_M1
         );
END_REGION

REGION Network 7: Activate cleaning piston mixinghead by external signal
         A     "DB005_RS<->Extern".MC_Interface[4].Data_from_MC.CP_forward;
         =     #Temp_CP_forward_external;
END_REGION

REGION Network 8: Cleaning piston mixinghead 04
         CALL  BLKMOV
         ( SRCBLK  := "DB123_MH_IO_Signals".MH[4].IN.CleaningPistonState,
           RET_VAL := #RetValSFC,
           DSTBLK  := #AnaCp_Stat
         );

         L     #AnaCp_Stat;
         SRW   8;
         T     #AnaCp_StatB;

         CALL  "FC071_CleaningPiston"
         ( IN_WithCP                := "DB704_MH_Value".Mixinghead[4].WithCleaningPiston,
           IN_Ana_CP_State          := #AnaCp_StatB,
           IN_SWUEnabled            := "DB619_State_MPart".SWU[1].SWU_released."04",
           IN_ButtonCPForward       := "DB123_MH_IO_Signals".MH[4].IN.MH_CP_forward,
           IN_ButtonCPback          := "DB123_MH_IO_Signals".MH[4].IN.MH_CP_backward,
           IN_CPForwardFromExternal := #Temp_CP_forward_external,
           IN_CPAfterShot           := "DB619_State_MPart".ShotMa[1].ShotData.CP_AfterShot,
           IN_PartshotDisabled      := "DB619_State_MPart".ShotMa[1].ShotData.ShotDisabled,
           IN_Blowing_OUT           := "DB614_MH_State".InertingMH[4].Start_Prepare_Purge_after_Shot,
           IN_CPProxSwitch          := "DB123_MH_IO_Signals".MH[4].IN.MH_APS_CleaningPiston,
           IN_SWUActive             := "DB619_State_MPart".SWU[1].Open_SWU_allone."04",
           IN_HydraulicOk           := "DB619_State_MPart".Machine[1].HydStartUp_finished,
           IN_ResetFaults           := "DB009_Faults".Faults_Reset_FKT_M1,
           IN_ControlVoltage        := "DB619_State_MPart".Operationmode[1].Controllvoltage,
           IN_OperatingModeValid    := "DB619_State_MPart".Operationmode[1].valid,
           IN_OperatingModeWithFoam := "DB619_State_MPart".Operationmode[1].Operation,
           IN_OperatingModeTestValv := "DB619_State_MPart".Operationmode[1].Test,
           IN_Lamptest              := "DB619_State_MPart".Operationmode[1].Lamptest,
           IN_ShotEnd               := "DB619_State_MPart".Cycle[1].PulsShotend,
           IN_FaultLevel_1          := "DB009_Faults".Fault_State_Grp_1_M1,
           IN_PressurizeTimeRunning := "DB619_State_MPart".Cycle[1].PressurizeTimeRuns,
           IN_ShotActive            := "DB619_State_MPart".Cycle[1].ShotRuns,
           IN_CycleRunning          := "DB619_State_MPart".Cycle[1].running,
           IN_RmpCtrlChangeTimeEnd  := "DB619_State_MPart".Cycle[1].RmpCtrlChangeTimeEnd,
           IN_StandbyTimeRunning    := "DB619_State_MPart".Cycle[1].StandByTimeRuns,
           IN_RmpCycleEnd           := "DB619_State_MPart".Cycle[1].PulseCycleEnd,
           IN_CPTimer               := "TM_RunTime_CP04",
           IN_TMCheckHomePos        := "TM_FltCPHomePos_CP04",
           Values                   := "DB704_MH_Value".Mixinghead[4].Cleaning_Piston,
           OUT_ValveCPForward       := "DB123_MH_IO_Signals".MH[4].OUT.MH.V_CP_Forward_MH,
           OUT_LampCPBack           := "DB123_MH_IO_Signals".MH[4].OUT.MH.H_CP_Back_MH,
           IO_CPIsOk                := "DB619_State_MPart".Mixinghead[1].Cleaningpiston_OK,
           IO_ReqHydrForCleaning    := "DB611_Hydraulic_State".MH_Hydraulic[1].Request_from_CP,
           IO_Status                := "DB614_MH_State".MH_CleaningPiston[4],
           IO_Fault                 := "DB824_Error_MH_CP".CPiston[4],
           IO_NewFault              := "DB009_Faults".Faultschanging_M1,
           IO_FaultLevel_1          := "DB009_Faults".Faults_FKT_Grp_1_M1,
           IO_FaultLevel_2          := "DB009_Faults".Faults_FKT_Grp_2_M1,
           IO_FaultLevel_3          := "DB009_Faults".Faults_FKT_Grp_3_M1
         );
END_REGION

REGION Network 9: Activate cleaning piston mixinghead by external signal
         A     "DB005_RS<->Extern".MC_Interface[5].Data_from_MC.CP_forward;
         =     #Temp_CP_forward_external;
END_REGION

REGION Network 10: Cleaning piston mixinghead 05
         CALL  BLKMOV
         ( SRCBLK  := "DB123_MH_IO_Signals".MH[5].IN.CleaningPistonState,
           RET_VAL := #RetValSFC,
           DSTBLK  := #AnaCp_Stat
         );

         L     #AnaCp_Stat;
         SRW   8;
         T     #AnaCp_StatB;

